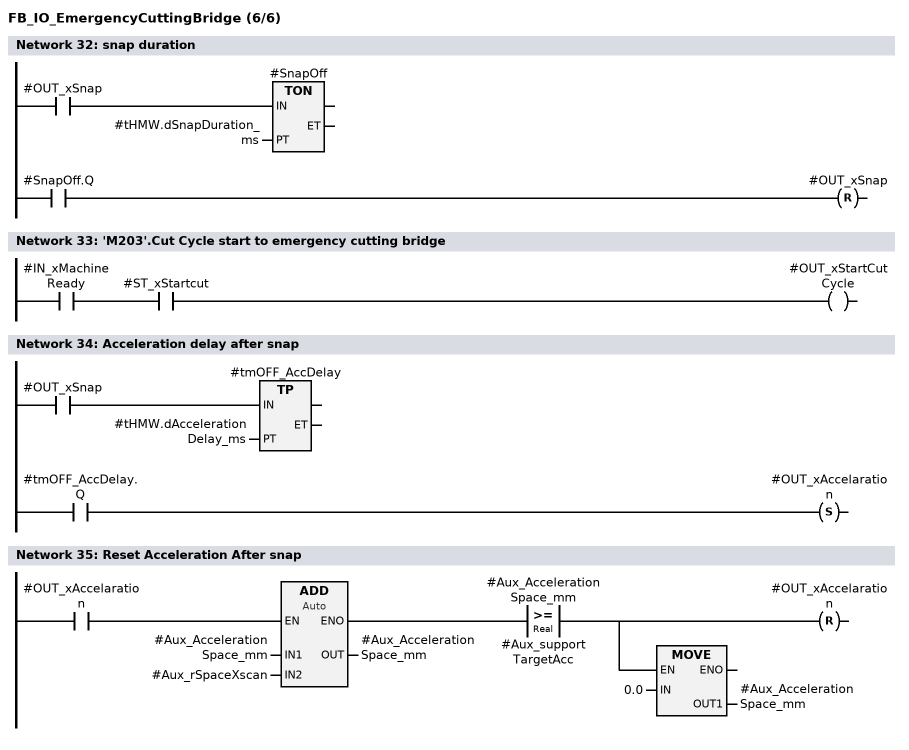
   #SnapOff(IN := #OUT_xSnap, PT := #tHMW.dSnapDuration_ms);   // TON
   IF #SnapOff.Q THEN #OUT_xSnap := FALSE; END_IF;
END_REGION

REGION Network 33: 'M203'.Cut Cycle start to emergency cutting bridge
   RUNG wire#powerrail
      Contact( #IN_xMachineReady )
      Contact( #ST_xStartcut )
      Coil( #OUT_xStartCutCycle )
   END_RUNG
   // the same network as SCL:
   #OUT_xStartCutCycle := #IN_xMachineReady AND #ST_xStartcut;
END_REGION

REGION Network 34: Acceleration delay after snap
   #tmOFF_AccDelay(IN := #OUT_xSnap, PT := #tHMW.dAccelerationDelay_ms);   // TP
   IF #tmOFF_AccDelay.Q THEN #OUT_xAccelaration := TRUE; END_IF;
END_REGION

REGION Network 35: Reset Acceleration After snap
   RUNG wire#powerrail
      Contact( #OUT_xAccelaration )
      Add(in1 := #Aux_AccelerationSpace_mm, in2 := #Aux_rSpaceXscan, out => #Aux_AccelerationSpace_mm)
      { S7_Templates := "SrcType := Real" } GE_Contact(in1 := #Aux_AccelerationSpace_mm, in2 := #Aux_supportTargetAcc)
      wire#w1
      R_Coil( #OUT_xAccelaration )
   END_RUNG
   RUNG wire#w1
      Move(in := 0.0, out1 => #Aux_AccelerationSpace_mm)
   END_RUNG
   // the same network as SCL:
   IF #OUT_xAccelaration THEN
       #Aux_AccelerationSpace_mm := #Aux_AccelerationSpace_mm + #Aux_rSpaceXscan;
   END_IF;
   #_w1 := #OUT_xAccelaration AND (#Aux_AccelerationSpace_mm >= #Aux_supportTargetAcc);
   IF #_w1 THEN
       #OUT_xAccelaration := FALSE;
       #Aux_AccelerationSpace_mm := 0.0;
   END_IF;
END_REGION
END_FUNCTION_BLOCK

// folder: 05_Reports

FUNCTION "RP_MergeToMergeMessageV2" : Void   // FC3, SCL
TITLE = RP_MergeMessage
{ S7_Optimized_Access := 'TRUE' }
AUTHOR : Cigliutt
FAMILY : RP
VERSION : 1.0
// This FC will be merge different flush buffer
   VAR_INPUT
      IN_xInit : Bool;   // Initialize the buffer container
   END_VAR
   VAR_IN_OUT
      INO_tMergeBuffer : "UDT_RP_MessageContMerge_v2";   // Merge buffer container
      INO_tMergeBuffer_1 : "UDT_RP_MessageContMerge_v2";   // Merge buffer container #1
      INO_tMergeBuffer_2 : "UDT_RP_MessageContMerge_v2";   // Merge buffer container #2
      INO_tMergeBuffer_3 : "UDT_RP_MessageContMerge_v2";   // Merge buffer container #3
      INO_tMergeBuffer_4 : "UDT_RP_MessageContMerge_v2";   // Merge buffer container #4
      INO_tMergeBuffer_5 : "UDT_RP_MessageContMerge_v2";   // Merge buffer container #5
      INO_xError : Bool;   // If =true error on flush
   END_VAR
   VAR_TEMP
      TMP_dIndex : DInt;
      TMP_dArrayNumEl : DInt;
      TMP_dtDateTime : Date_And_Time;
      TMP_dRetVal : DInt;
      TMP_dDataToCopy : DInt;
      TMP_dOldNumMex : DInt;
      TMP_dActualNumMex : DInt;
   END_VAR
BEGIN
   //Manage the initialization request. Fill to 0 the buffer and the values.
   //After that calculate the space available
   //
   #TMP_dRetVal := RD_LOC_T(#TMP_dtDateTime);

   IF #IN_xInit = true THEN

       //Initialize the values
       #INO_tMergeBuffer.dNumOfMessage := 0;
       #INO_tMergeBuffer.dMaxNumOfMessage := 0;

       //Take the number OF elements OF the array data, reset it AND set the number
       //to iDataMaxElem
       #TMP_dArrayNumEl := "GP_GetArraySize"(INO_vArray := #INO_tMergeBuffer.rgtMessages);

       #INO_tMergeBuffer.dMaxNumOfMessage := #TMP_dArrayNumEl;

       //Reset the buffer
       //

       FOR #TMP_dIndex := 0 TO #INO_tMergeBuffer.dMaxNumOfMessage - 1 DO
           #INO_tMergeBuffer.rgtMessages[#TMP_dIndex].dCodeEvent := 0;
           #INO_tMergeBuffer.rgtMessages[#TMP_dIndex].dEvent1 := 0;
           #INO_tMergeBuffer.rgtMessages[#TMP_dIndex].dEvent2 := 0;
           #INO_tMergeBuffer.rgtMessages[#TMP_dIndex].dEvent3 := 0;
           #INO_tMergeBuffer.rgtMessages[#TMP_dIndex].dEvent4 := 0;
           #INO_tMergeBuffer.rgtMessages[#TMP_dIndex].dEvent5 := 0;
           #INO_tMergeBuffer.rgtMessages[#TMP_dIndex].dEvent6 := 0;
           #INO_tMergeBuffer.rgtMessages[#TMP_dIndex].dEvent7 := 0;
           #INO_tMergeBuffer.rgtMessages[#TMP_dIndex].dEvent8 := 0;
           #INO_tMergeBuffer.rgtMessages[#TMP_dIndex].dEvent9 := 0;
           #INO_tMergeBuffer.rgtMessages[#TMP_dIndex].dEvent10 := 0;

           #INO_tMergeBuffer.rgtMessages[#TMP_dIndex].strIdent := '';
           #INO_tMergeBuffer.rgtMessages[#TMP_dIndex].dtDateTime := #TMP_dtDateTime;
       END_FOR;

       #INO_tMergeBuffer.xInitialized := true;

       RETURN;
   END_IF;

   //If we are not in initializing mode, copy the input value inside the array.
   //First of all check if the data are consistent
   //
   IF (#INO_tMergeBuffer.xInitialized = false) OR
       (#INO_tMergeBuffer_1.xInitialized = false) OR
       (#INO_tMergeBuffer_2.xInitialized = false) OR
       (#INO_tMergeBuffer_3.xInitialized = false) OR
       (#INO_tMergeBuffer_4.xInitialized = false) OR
       (#INO_tMergeBuffer_5.xInitialized = false) THEN

       #INO_xError := true;

       RETURN;
   END_IF;

   //Check if the merge buffer is free. Otherwise exit
   //
   IF (#INO_tMergeBuffer.dNumOfMessage > 0) THEN
       RETURN;
   END_IF;


   ///*********************************** FLUSH BUFFER #1

   //Check if the first flush buffer, has data inside
   IF (#INO_tMergeBuffer_1.dNumOfMessage > 0) THEN

       #TMP_dDataToCopy := #INO_tMergeBuffer_1.dNumOfMessage;

       IF (#TMP_dDataToCopy > #INO_tMergeBuffer.dMaxNumOfMessage) THEN
           #TMP_dDataToCopy := #INO_tMergeBuffer.dMaxNumOfMessage;
       END_IF;

       //Copy the data
       #TMP_dRetVal := "GP_BlockMoveStruct"(IN_iSourceIndex := 0,
                                            IN_iDestIndex := 0,
                                            IN_iCount := DINT_TO_INT(#TMP_dDataToCopy),
                                            INO_vSourceArrayStruct := #INO_tMergeBuffer_1.rgtMessages,
                                            INO_vDestArrayStruct := #INO_tMergeBuffer.rgtMessages);

       #INO_tMergeBuffer.dNumOfMessage := #TMP_dDataToCopy;

       //Check if some data is remaining. If yes, compact it on the FlushBuffer
       //
       IF (#INO_tMergeBuffer_1.dNumOfMessage - #TMP_dDataToCopy) > 0 THEN
           //Copy the data
           #TMP_dRetVal := "GP_BlockMoveStruct"(IN_iSourceIndex := DINT_TO_INT(#INO_tMergeBuffer_1.dNumOfMessage - (#INO_tMergeBuffer_1.dNumOfMessage - #TMP_dDataToCopy)),
                                                IN_iDestIndex := 0,
                                                IN_iCount := DINT_TO_INT(#INO_tMergeBuffer_1.dNumOfMessage - #TMP_dDataToCopy),
                                                INO_vSourceArrayStruct := #INO_tMergeBuffer_1.rgtMessages,
                                                INO_vDestArrayStruct := #INO_tMergeBuffer_1.rgtMessages);


       END_IF;

       #TMP_dOldNumMex := #INO_tMergeBuffer_1.dNumOfMessage;
       #TMP_dActualNumMex := #INO_tMergeBuffer_1.dNumOfMessage - #TMP_dDataToCopy;


       //Data moved, fill the remaining buffer. To increase performance, fill only the data that was used
       //
       FOR #TMP_dIndex := #TMP_dActualNumMex TO #TMP_dOldNumMex - 1 DO

           #INO_tMergeBuffer_1.rgtMessages[#TMP_dIndex].dCodeEvent := 0;
           #INO_tMergeBuffer_1.rgtMessages[#TMP_dIndex].dEvent1 := 0;
           #INO_tMergeBuffer_1.rgtMessages[#TMP_dIndex].dEvent2 := 0;
           #INO_tMergeBuffer_1.rgtMessages[#TMP_dIndex].dEvent3 := 0;
           #INO_tMergeBuffer_1.rgtMessages[#TMP_dIndex].dEvent4 := 0;
           #INO_tMergeBuffer_1.rgtMessages[#TMP_dIndex].dEvent5 := 0;
           #INO_tMergeBuffer_1.rgtMessages[#TMP_dIndex].dEvent6 := 0;
           #INO_tMergeBuffer_1.rgtMessages[#TMP_dIndex].dEvent7 := 0;
           #INO_tMergeBuffer_1.rgtMessages[#TMP_dIndex].dEvent8 := 0;
           #INO_tMergeBuffer_1.rgtMessages[#TMP_dIndex].dEvent9 := 0;
           #INO_tMergeBuffer_1.rgtMessages[#TMP_dIndex].dEvent10 := 0;

           #INO_tMergeBuffer_1.rgtMessages[#TMP_dIndex].strIdent := '';
           #INO_tMergeBuffer_1.rgtMessages[#TMP_dIndex].dtDateTime := #TMP_dtDateTime;
       END_FOR;

       #INO_tMergeBuffer_1.dNumOfMessage := #TMP_dActualNumMex;

   END_IF;


   ///*********************************** FLUSH BUFFER #2

   //Check if the first flush buffer, has data inside
   IF (#INO_tMergeBuffer_2.dNumOfMessage > 0) AND (#INO_tMergeBuffer.dNumOfMessage < #INO_tMergeBuffer.dMaxNumOfMessage) THEN

       #TMP_dDataToCopy := #INO_tMergeBuffer_2.dNumOfMessage;

       IF (#TMP_dDataToCopy + #INO_tMergeBuffer.dNumOfMessage > #INO_tMergeBuffer.dMaxNumOfMessage) THEN
           #TMP_dDataToCopy := #INO_tMergeBuffer.dMaxNumOfMessage - #INO_tMergeBuffer.dNumOfMessage;
       END_IF;

       //Copy the data
       #TMP_dRetVal := "GP_BlockMoveStruct"(IN_iSourceIndex := 0,
                                            IN_iDestIndex := DINT_TO_INT(#INO_tMergeBuffer.dNumOfMessage),
                                            IN_iCount := DINT_TO_INT(#TMP_dDataToCopy),
                                            INO_vSourceArrayStruct := #INO_tMergeBuffer_2.rgtMessages,
                                            INO_vDestArrayStruct := #INO_tMergeBuffer.rgtMessages);

       #INO_tMergeBuffer.dNumOfMessage := #INO_tMergeBuffer.dNumOfMessage + #TMP_dDataToCopy;

       //Check if some data is remaining. If yes, compact it on the FlushBuffer
       //
       IF (#INO_tMergeBuffer_2.dNumOfMessage - #TMP_dDataToCopy) > 0 THEN
           //Copy the data
           #TMP_dRetVal := "GP_BlockMoveStruct"(IN_iSourceIndex := DINT_TO_INT(#INO_tMergeBuffer_2.dNumOfMessage - (#INO_tMergeBuffer_2.dNumOfMessage - #TMP_dDataToCopy)),
                                                IN_iDestIndex := 0,
                                                IN_iCount := DINT_TO_INT(#INO_tMergeBuffer_2.dNumOfMessage - #TMP_dDataToCopy),
                                                INO_vSourceArrayStruct := #INO_tMergeBuffer_2.rgtMessages,
                                                INO_vDestArrayStruct := #INO_tMergeBuffer_2.rgtMessages);


       END_IF;

       #TMP_dOldNumMex := #INO_tMergeBuffer_2.dNumOfMessage;
       #TMP_dActualNumMex := #INO_tMergeBuffer_2.dNumOfMessage - #TMP_dDataToCopy;



       //Data moved, fill the remaining buffer. To increase performance, fill only the data that was used
       //
       FOR #TMP_dIndex := #TMP_dActualNumMex TO #TMP_dOldNumMex - 1 DO

           #INO_tMergeBuffer_2.rgtMessages[#TMP_dIndex].dCodeEvent := 0;
           #INO_tMergeBuffer_2.rgtMessages[#TMP_dIndex].dEvent1 := 0;
           #INO_tMergeBuffer_2.rgtMessages[#TMP_dIndex].dEvent2 := 0;
           #INO_tMergeBuffer_2.rgtMessages[#TMP_dIndex].dEvent3 := 0;
           #INO_tMergeBuffer_2.rgtMessages[#TMP_dIndex].dEvent4 := 0;
           #INO_tMergeBuffer_2.rgtMessages[#TMP_dIndex].dEvent5 := 0;
           #INO_tMergeBuffer_2.rgtMessages[#TMP_dIndex].dEvent6 := 0;
           #INO_tMergeBuffer_2.rgtMessages[#TMP_dIndex].dEvent7 := 0;
           #INO_tMergeBuffer_2.rgtMessages[#TMP_dIndex].dEvent8 := 0;
           #INO_tMergeBuffer_2.rgtMessages[#TMP_dIndex].dEvent9 := 0;
           #INO_tMergeBuffer_2.rgtMessages[#TMP_dIndex].dEvent10 := 0;
           #INO_tMergeBuffer_2.rgtMessages[#TMP_dIndex].strIdent := '';

           #INO_tMergeBuffer_2.rgtMessages[#TMP_dIndex].dtDateTime := #TMP_dtDateTime;
       END_FOR;

       #INO_tMergeBuffer_2.dNumOfMessage := #TMP_dActualNumMex;
   END_IF;


   ///*********************************** FLUSH BUFFER #3


   //Check if the first flush buffer, has data inside
   IF (#INO_tMergeBuffer_3.dNumOfMessage > 0) AND (#INO_tMergeBuffer.dNumOfMessage < #INO_tMergeBuffer.dMaxNumOfMessage) THEN

       #TMP_dDataToCopy := #INO_tMergeBuffer_3.dNumOfMessage;

       IF (#TMP_dDataToCopy + #INO_tMergeBuffer.dNumOfMessage > #INO_tMergeBuffer.dMaxNumOfMessage) THEN
           #TMP_dDataToCopy := #INO_tMergeBuffer.dMaxNumOfMessage - #INO_tMergeBuffer.dNumOfMessage;
       END_IF;

       //Copy the data
       #TMP_dRetVal := "GP_BlockMoveStruct"(IN_iSourceIndex := 0,
                                            IN_iDestIndex := DINT_TO_INT(#INO_tMergeBuffer.dNumOfMessage),
                                            IN_iCount := DINT_TO_INT(#TMP_dDataToCopy),
                                            INO_vSourceArrayStruct := #INO_tMergeBuffer_3.rgtMessages,
                                            INO_vDestArrayStruct := #INO_tMergeBuffer.rgtMessages);

       #INO_tMergeBuffer.dNumOfMessage := #INO_tMergeBuffer.dNumOfMessage + #TMP_dDataToCopy;

       //Check if some data is remaining. If yes, compact it on the FlushBuffer
       //
       IF (#INO_tMergeBuffer_3.dNumOfMessage - #TMP_dDataToCopy) > 0 THEN
           //Copy the data
           #TMP_dRetVal := "GP_BlockMoveStruct"(IN_iSourceIndex := DINT_TO_INT(#INO_tMergeBuffer_3.dNumOfMessage - (#INO_tMergeBuffer_3.dNumOfMessage - #TMP_dDataToCopy)),
                                                IN_iDestIndex := 0,
                                                IN_iCount := DINT_TO_INT(#INO_tMergeBuffer_3.dNumOfMessage - #TMP_dDataToCopy),
                                                INO_vSourceArrayStruct := #INO_tMergeBuffer_3.rgtMessages,
                                                INO_vDestArrayStruct := #INO_tMergeBuffer_3.rgtMessages);


       END_IF;

       #TMP_dOldNumMex := #INO_tMergeBuffer_3.dNumOfMessage;
       #TMP_dActualNumMex := #INO_tMergeBuffer_3.dNumOfMessage - #TMP_dDataToCopy;


       //Data moved, fill the remaining buffer. To increase performance, fill only the data that was used
       //
       FOR #TMP_dIndex := #TMP_dActualNumMex TO #TMP_dOldNumMex - 1 DO

           #INO_tMergeBuffer_3.rgtMessages[#TMP_dIndex].dCodeEvent := 0;
           #INO_tMergeBuffer_3.rgtMessages[#TMP_dIndex].dEvent1 := 0;
           #INO_tMergeBuffer_3.rgtMessages[#TMP_dIndex].dEvent2 := 0;
           #INO_tMergeBuffer_3.rgtMessages[#TMP_dIndex].dEvent3 := 0;
           #INO_tMergeBuffer_3.rgtMessages[#TMP_dIndex].dEvent4 := 0;
           #INO_tMergeBuffer_3.rgtMessages[#TMP_dIndex].dEvent5 := 0;
           #INO_tMergeBuffer_3.rgtMessages[#TMP_dIndex].dEvent6 := 0;
           #INO_tMergeBuffer_3.rgtMessages[#TMP_dIndex].dEvent7 := 0;
           #INO_tMergeBuffer_3.rgtMessages[#TMP_dIndex].dEvent8 := 0;
           #INO_tMergeBuffer_3.rgtMessages[#TMP_dIndex].dEvent9 := 0;
           #INO_tMergeBuffer_3.rgtMessages[#TMP_dIndex].dEvent10 := 0;
           #INO_tMergeBuffer_3.rgtMessages[#TMP_dIndex].strIdent := '';

           #INO_tMergeBuffer_3.rgtMessages[#TMP_dIndex].dtDateTime := #TMP_dtDateTime;
       END_FOR;

       #INO_tMergeBuffer_3.dNumOfMessage := #TMP_dActualNumMex;


   END_IF;


   ///*********************************** FLUSH BUFFER #4


   //Check if the first flush buffer, has data inside
   IF (#INO_tMergeBuffer_4.dNumOfMessage > 0) AND (#INO_tMergeBuffer.dNumOfMessage < #INO_tMergeBuffer.dMaxNumOfMessage) THEN

       #TMP_dDataToCopy := #INO_tMergeBuffer_4.dNumOfMessage;

       IF (#TMP_dDataToCopy + #INO_tMergeBuffer.dNumOfMessage > #INO_tMergeBuffer.dMaxNumOfMessage) THEN
           #TMP_dDataToCopy := #INO_tMergeBuffer.dMaxNumOfMessage - #INO_tMergeBuffer.dNumOfMessage;
       END_IF;

       //Copy the data
       #TMP_dRetVal := "GP_BlockMoveStruct"(IN_iSourceIndex := 0,
                                            IN_iDestIndex := DINT_TO_INT(#INO_tMergeBuffer.dNumOfMessage),
                                            IN_iCount := DINT_TO_INT(#TMP_dDataToCopy),
                                            INO_vSourceArrayStruct := #INO_tMergeBuffer_4.rgtMessages,
                                            INO_vDestArrayStruct := #INO_tMergeBuffer.rgtMessages);

       #INO_tMergeBuffer.dNumOfMessage := #INO_tMergeBuffer.dNumOfMessage + #TMP_dDataToCopy;

       //Check if some data is remaining. If yes, compact it on the FlushBuffer
       //
       IF (#INO_tMergeBuffer_4.dNumOfMessage - #TMP_dDataToCopy) > 0 THEN
           //Copy the data
           #TMP_dRetVal := "GP_BlockMoveStruct"(IN_iSourceIndex := DINT_TO_INT(#INO_tMergeBuffer_4.dNumOfMessage - (#INO_tMergeBuffer_4.dNumOfMessage - #TMP_dDataToCopy)),
                                                IN_iDestIndex := 0,
                                                IN_iCount := DINT_TO_INT(#INO_tMergeBuffer_4.dNumOfMessage - #TMP_dDataToCopy),
                                                INO_vSourceArrayStruct := #INO_tMergeBuffer_4.rgtMessages,
                                                INO_vDestArrayStruct := #INO_tMergeBuffer_4.rgtMessages);


       END_IF;

       #TMP_dOldNumMex := #INO_tMergeBuffer_4.dNumOfMessage;
       #TMP_dActualNumMex := #INO_tMergeBuffer_4.dNumOfMessage - #TMP_dDataToCopy;


       //Data moved, fill the remaining buffer. To increase performance, fill only the data that was used
       //
       FOR #TMP_dIndex := #TMP_dActualNumMex TO #TMP_dOldNumMex - 1 DO

           #INO_tMergeBuffer_4.rgtMessages[#TMP_dIndex].dCodeEvent := 0;
           #INO_tMergeBuffer_4.rgtMessages[#TMP_dIndex].dEvent1 := 0;
           #INO_tMergeBuffer_4.rgtMessages[#TMP_dIndex].dEvent2 := 0;
           #INO_tMergeBuffer_4.rgtMessages[#TMP_dIndex].dEvent3 := 0;
           #INO_tMergeBuffer_4.rgtMessages[#TMP_dIndex].dEvent4 := 0;
           #INO_tMergeBuffer_4.rgtMessages[#TMP_dIndex].dEvent5 := 0;
           #INO_tMergeBuffer_4.rgtMessages[#TMP_dIndex].dEvent6 := 0;
           #INO_tMergeBuffer_4.rgtMessages[#TMP_dIndex].dEvent7 := 0;
           #INO_tMergeBuffer_4.rgtMessages[#TMP_dIndex].dEvent8 := 0;
           #INO_tMergeBuffer_4.rgtMessages[#TMP_dIndex].dEvent9 := 0;
           #INO_tMergeBuffer_4.rgtMessages[#TMP_dIndex].dEvent10 := 0;
           #INO_tMergeBuffer_4.rgtMessages[#TMP_dIndex].strIdent := '';

           #INO_tMergeBuffer_4.rgtMessages[#TMP_dIndex].dtDateTime := #TMP_dtDateTime;
       END_FOR;

       #INO_tMergeBuffer_4.dNumOfMessage := #TMP_dActualNumMex;


   END_IF;


   ///*********************************** FLUSH BUFFER #5


   //Check if the first flush buffer, has data inside
   IF (#INO_tMergeBuffer_5.dNumOfMessage > 0) AND (#INO_tMergeBuffer.dNumOfMessage < #INO_tMergeBuffer.dMaxNumOfMessage) THEN

       #TMP_dDataToCopy := #INO_tMergeBuffer_5.dNumOfMessage;

       IF (#TMP_dDataToCopy + #INO_tMergeBuffer.dNumOfMessage > #INO_tMergeBuffer.dMaxNumOfMessage) THEN
           #TMP_dDataToCopy := #INO_tMergeBuffer.dMaxNumOfMessage - #INO_tMergeBuffer.dNumOfMessage;
       END_IF;

       //Copy the data
       #TMP_dRetVal := "GP_BlockMoveStruct"(IN_iSourceIndex := 0,
                                            IN_iDestIndex := DINT_TO_INT(#INO_tMergeBuffer.dNumOfMessage),
                                            IN_iCount := DINT_TO_INT(#TMP_dDataToCopy),
                                            INO_vSourceArrayStruct := #INO_tMergeBuffer_5.rgtMessages,
                                            INO_vDestArrayStruct := #INO_tMergeBuffer.rgtMessages);

       #INO_tMergeBuffer.dNumOfMessage := #INO_tMergeBuffer.dNumOfMessage + #TMP_dDataToCopy;

       //Check if some data is remaining. If yes, compact it on the FlushBuffer
       //
       IF (#INO_tMergeBuffer_5.dNumOfMessage - #TMP_dDataToCopy) > 0 THEN
           //Copy the data
           #TMP_dRetVal := "GP_BlockMoveStruct"(IN_iSourceIndex := DINT_TO_INT(#INO_tMergeBuffer_5.dNumOfMessage - (#INO_tMergeBuffer_5.dNumOfMessage - #TMP_dDataToCopy)),
                                                IN_iDestIndex := 0,
                                                IN_iCount := DINT_TO_INT(#INO_tMergeBuffer_5.dNumOfMessage - #TMP_dDataToCopy),
                                                INO_vSourceArrayStruct := #INO_tMergeBuffer_5.rgtMessages,
                                                INO_vDestArrayStruct := #INO_tMergeBuffer_5.rgtMessages);


       END_IF;

       #TMP_dOldNumMex := #INO_tMergeBuffer_5.dNumOfMessage;
       #TMP_dActualNumMex := #INO_tMergeBuffer_5.dNumOfMessage - #TMP_dDataToCopy;

       //Data moved, fill the remaining buffer. To increase performance, fill only the data that was used
       //
       FOR #TMP_dIndex := #TMP_dActualNumMex TO #TMP_dOldNumMex - 1 DO

           #INO_tMergeBuffer_5.rgtMessages[#TMP_dIndex].dCodeEvent := 0;
           #INO_tMergeBuffer_5.rgtMessages[#TMP_dIndex].dEvent1 := 0;
           #INO_tMergeBuffer_5.rgtMessages[#TMP_dIndex].dEvent2 := 0;
           #INO_tMergeBuffer_5.rgtMessages[#TMP_dIndex].dEvent3 := 0;
           #INO_tMergeBuffer_5.rgtMessages[#TMP_dIndex].dEvent4 := 0;
           #INO_tMergeBuffer_5.rgtMessages[#TMP_dIndex].dEvent5 := 0;
           #INO_tMergeBuffer_5.rgtMessages[#TMP_dIndex].dEvent6 := 0;
           #INO_tMergeBuffer_5.rgtMessages[#TMP_dIndex].dEvent7 := 0;
           #INO_tMergeBuffer_5.rgtMessages[#TMP_dIndex].dEvent8 := 0;
           #INO_tMergeBuffer_5.rgtMessages[#TMP_dIndex].dEvent9 := 0;
           #INO_tMergeBuffer_5.rgtMessages[#TMP_dIndex].dEvent10 := 0;
           #INO_tMergeBuffer_5.rgtMessages[#TMP_dIndex].strIdent := '';

           #INO_tMergeBuffer_5.rgtMessages[#TMP_dIndex].dtDateTime := #TMP_dtDateTime;
       END_FOR;

       #INO_tMergeBuffer_5.dNumOfMessage := #TMP_dActualNumMex;


   END_IF;
END_FUNCTION

FUNCTION "RP_OB_TaskSlowToOpt" : Void   // FC4, LAD
{ S7_Optimized_Access := 'TRUE' }
VERSION : 0.1
   VAR_INPUT
      IN_xFirstScan : Bool;
   END_VAR
   VAR_TEMP
      TMP_xError : Bool;
   END_VAR
BEGIN

REGION Network 1
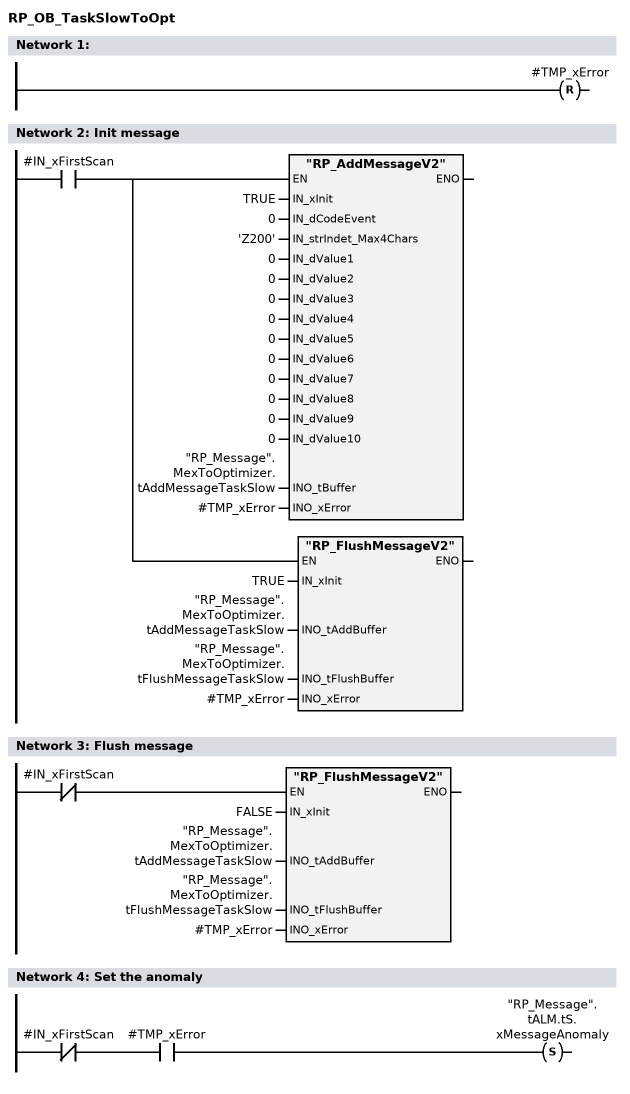
   RUNG wire#powerrail
      R_Coil( #TMP_xError )
   END_RUNG
   // the same network as SCL:
   #TMP_xError := FALSE;
END_REGION

REGION Network 2: Init message
   RUNG wire#powerrail
      Contact( #IN_xFirstScan )
      wire#w1
      "RP_AddMessageV2"(IN_xInit := TRUE, IN_dCodeEvent := 0, IN_strIndet_Max4Chars := 'Z200', IN_dValue1 := 0, IN_dValue2 := 0, IN_dValue3 := 0, IN_dValue4 := 0, IN_dValue5 := 0, IN_dValue6 := 0, IN_dValue7 := 0, IN_dValue8 := 0, IN_dValue9 := 0, IN_dValue10 := 0, INO_tBuffer := "RP_Message".MexToOptimizer.tAddMessageTaskSlow, INO_xError := #TMP_xError)
   END_RUNG
   RUNG wire#w1
      "RP_FlushMessageV2"(IN_xInit := TRUE, INO_tAddBuffer := "RP_Message".MexToOptimizer.tAddMessageTaskSlow, INO_tFlushBuffer := "RP_Message".MexToOptimizer.tFlushMessageTaskSlow, INO_xError := #TMP_xError)
   END_RUNG
   // the same network as SCL:
   IF #IN_xFirstScan THEN
       "RP_AddMessageV2"(IN_xInit := TRUE,
                         IN_dCodeEvent := 0,
                         IN_strIndet_Max4Chars := 'Z200',
                         IN_dValue1 := 0,
                         IN_dValue2 := 0,
                         IN_dValue3 := 0,
                         IN_dValue4 := 0,
                         IN_dValue5 := 0,
                         IN_dValue6 := 0,
                         IN_dValue7 := 0,
                         IN_dValue8 := 0,
                         IN_dValue9 := 0,
                         IN_dValue10 := 0,
                         INO_tBuffer := "RP_Message".MexToOptimizer.tAddMessageTaskSlow,
                         INO_xError := #TMP_xError);
       "RP_FlushMessageV2"(IN_xInit := TRUE,
                           INO_tAddBuffer := "RP_Message".MexToOptimizer.tAddMessageTaskSlow,
                           INO_tFlushBuffer := "RP_Message".MexToOptimizer.tFlushMessageTaskSlow,
                           INO_xError := #TMP_xError);
   END_IF;
END_REGION

REGION Network 3: Flush message
   RUNG wire#powerrail
      I_Contact( #IN_xFirstScan )
      "RP_FlushMessageV2"(IN_xInit := FALSE, INO_tAddBuffer := "RP_Message".MexToOptimizer.tAddMessageTaskSlow, INO_tFlushBuffer := "RP_Message".MexToOptimizer.tFlushMessageTaskSlow, INO_xError := #TMP_xError)
   END_RUNG
   // the same network as SCL:
   IF NOT #IN_xFirstScan THEN
       "RP_FlushMessageV2"(IN_xInit := FALSE,
                           INO_tAddBuffer := "RP_Message".MexToOptimizer.tAddMessageTaskSlow,
                           INO_tFlushBuffer := "RP_Message".MexToOptimizer.tFlushMessageTaskSlow,
                           INO_xError := #TMP_xError);
   END_IF;
END_REGION

REGION Network 4: Set the anomaly
   RUNG wire#powerrail
      I_Contact( #IN_xFirstScan )
      Contact( #TMP_xError )
      S_Coil( "RP_Message".tALM.tS.xMessageAnomaly )
   END_RUNG
   // the same network as SCL:
   IF NOT #IN_xFirstScan AND #TMP_xError THEN "RP_Message".tALM.tS.xMessageAnomaly := TRUE; END_IF;
END_REGION
END_FUNCTION

FUNCTION "RP_OB_TaskMediumFromOpt" : Void   // FC5, LAD
{ S7_Optimized_Access := 'TRUE' }
VERSION : 0.1
   VAR_INPUT
      IN_xFirstScan : Bool;
   END_VAR
   VAR_TEMP
      TMP_xError : Bool;
   END_VAR
BEGIN

REGION Network 1
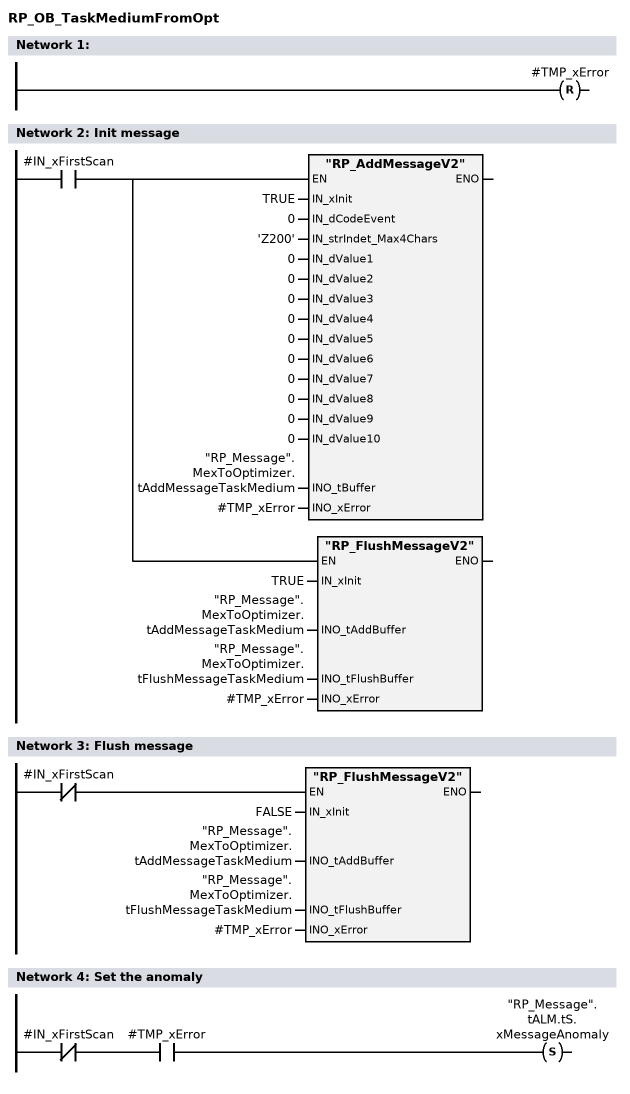
   RUNG wire#powerrail
      R_Coil( #TMP_xError )
   END_RUNG
   // the same network as SCL:
   #TMP_xError := FALSE;
END_REGION

REGION Network 2: Init message
   RUNG wire#powerrail
      Contact( #IN_xFirstScan )
      wire#w1
      "RP_AddMessageV2"(IN_xInit := TRUE, IN_dCodeEvent := 0, IN_strIndet_Max4Chars := 'Z200', IN_dValue1 := 0, IN_dValue2 := 0, IN_dValue3 := 0, IN_dValue4 := 0, IN_dValue5 := 0, IN_dValue6 := 0, IN_dValue7 := 0, IN_dValue8 := 0, IN_dValue9 := 0, IN_dValue10 := 0, INO_tBuffer := "RP_Message".MexToOptimizer.tAddMessageTaskMedium, INO_xError := #TMP_xError)
   END_RUNG
   RUNG wire#w1
      "RP_FlushMessageV2"(IN_xInit := TRUE, INO_tAddBuffer := "RP_Message".MexToOptimizer.tAddMessageTaskMedium, INO_tFlushBuffer := "RP_Message".MexToOptimizer.tFlushMessageTaskMedium, INO_xError := #TMP_xError)
   END_RUNG
   // the same network as SCL:
   IF #IN_xFirstScan THEN
       "RP_AddMessageV2"(IN_xInit := TRUE,
                         IN_dCodeEvent := 0,
                         IN_strIndet_Max4Chars := 'Z200',
                         IN_dValue1 := 0,
                         IN_dValue2 := 0,
                         IN_dValue3 := 0,
                         IN_dValue4 := 0,
                         IN_dValue5 := 0,
                         IN_dValue6 := 0,
                         IN_dValue7 := 0,
                         IN_dValue8 := 0,
                         IN_dValue9 := 0,
                         IN_dValue10 := 0,
                         INO_tBuffer := "RP_Message".MexToOptimizer.tAddMessageTaskMedium,
                         INO_xError := #TMP_xError);
       "RP_FlushMessageV2"(IN_xInit := TRUE,
                           INO_tAddBuffer := "RP_Message".MexToOptimizer.tAddMessageTaskMedium,
                           INO_tFlushBuffer := "RP_Message".MexToOptimizer.tFlushMessageTaskMedium,
                           INO_xError := #TMP_xError);
   END_IF;
END_REGION

REGION Network 3: Flush message
   RUNG wire#powerrail
      I_Contact( #IN_xFirstScan )
      "RP_FlushMessageV2"(IN_xInit := FALSE, INO_tAddBuffer := "RP_Message".MexToOptimizer.tAddMessageTaskMedium, INO_tFlushBuffer := "RP_Message".MexToOptimizer.tFlushMessageTaskMedium, INO_xError := #TMP_xError)
   END_RUNG
   // the same network as SCL:
   IF NOT #IN_xFirstScan THEN
       "RP_FlushMessageV2"(IN_xInit := FALSE,
                           INO_tAddBuffer := "RP_Message".MexToOptimizer.tAddMessageTaskMedium,
                           INO_tFlushBuffer := "RP_Message".MexToOptimizer.tFlushMessageTaskMedium,
                           INO_xError := #TMP_xError);
   END_IF;
END_REGION

REGION Network 4: Set the anomaly
   RUNG wire#powerrail
      I_Contact( #IN_xFirstScan )
      Contact( #TMP_xError )
      S_Coil( "RP_Message".tALM.tS.xMessageAnomaly )
   END_RUNG
   // the same network as SCL:
   IF NOT #IN_xFirstScan AND #TMP_xError THEN "RP_Message".tALM.tS.xMessageAnomaly := TRUE; END_IF;
END_REGION
END_FUNCTION

FUNCTION "RP_OB_TaskMediumToOpt" : Void   // FC6, LAD
{ S7_Optimized_Access := 'TRUE' }
VERSION : 0.1
   VAR_INPUT
      IN_xFirstScan : Bool;
   END_VAR
   VAR_TEMP
      TMP_xError : Bool;
   END_VAR
BEGIN

REGION Network 1
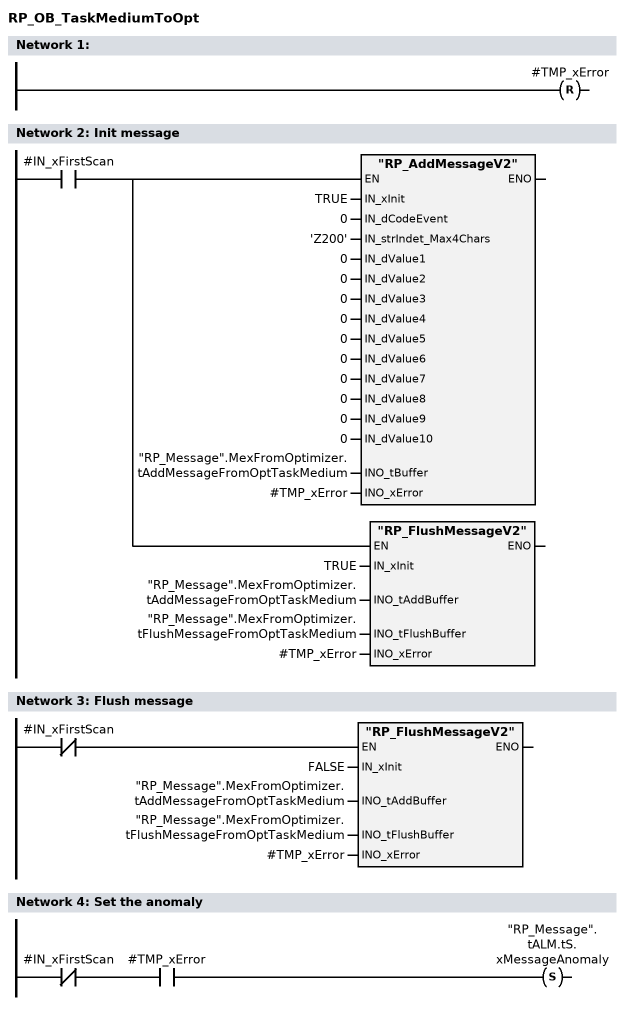
   RUNG wire#powerrail
      R_Coil( #TMP_xError )
   END_RUNG
   // the same network as SCL:
   #TMP_xError := FALSE;
END_REGION

REGION Network 2: Init message
   RUNG wire#powerrail
      Contact( #IN_xFirstScan )
      wire#w1
      "RP_AddMessageV2"(IN_xInit := TRUE, IN_dCodeEvent := 0, IN_strIndet_Max4Chars := 'Z200', IN_dValue1 := 0, IN_dValue2 := 0, IN_dValue3 := 0, IN_dValue4 := 0, IN_dValue5 := 0, IN_dValue6 := 0, IN_dValue7 := 0, IN_dValue8 := 0, IN_dValue9 := 0, IN_dValue10 := 0, INO_tBuffer := "RP_Message".MexFromOptimizer.tAddMessageFromOptTaskMedium, INO_xError := #TMP_xError)
   END_RUNG
   RUNG wire#w1
      "RP_FlushMessageV2"(IN_xInit := TRUE, INO_tAddBuffer := "RP_Message".MexFromOptimizer.tAddMessageFromOptTaskMedium, INO_tFlushBuffer := "RP_Message".MexFromOptimizer.tFlushMessageFromOptTaskMedium, INO_xError := #TMP_xError)
   END_RUNG
   // the same network as SCL:
   IF #IN_xFirstScan THEN
       "RP_AddMessageV2"(IN_xInit := TRUE,
                         IN_dCodeEvent := 0,
                         IN_strIndet_Max4Chars := 'Z200',
                         IN_dValue1 := 0,
                         IN_dValue2 := 0,
                         IN_dValue3 := 0,
                         IN_dValue4 := 0,
                         IN_dValue5 := 0,
                         IN_dValue6 := 0,
                         IN_dValue7 := 0,
                         IN_dValue8 := 0,
                         IN_dValue9 := 0,
                         IN_dValue10 := 0,
                         INO_tBuffer := "RP_Message".MexFromOptimizer.tAddMessageFromOptTaskMedium,
                         INO_xError := #TMP_xError);
       "RP_FlushMessageV2"(IN_xInit := TRUE,
                           INO_tAddBuffer := "RP_Message".MexFromOptimizer.tAddMessageFromOptTaskMedium,
                           INO_tFlushBuffer := "RP_Message".MexFromOptimizer.tFlushMessageFromOptTaskMedium,
                           INO_xError := #TMP_xError);
   END_IF;
END_REGION

REGION Network 3: Flush message
   RUNG wire#powerrail
      I_Contact( #IN_xFirstScan )
      "RP_FlushMessageV2"(IN_xInit := FALSE, INO_tAddBuffer := "RP_Message".MexFromOptimizer.tAddMessageFromOptTaskMedium, INO_tFlushBuffer := "RP_Message".MexFromOptimizer.tFlushMessageFromOptTaskMedium, INO_xError := #TMP_xError)
   END_RUNG
   // the same network as SCL:
   IF NOT #IN_xFirstScan THEN
       "RP_FlushMessageV2"(IN_xInit := FALSE,
                           INO_tAddBuffer := "RP_Message".MexFromOptimizer.tAddMessageFromOptTaskMedium,
                           INO_tFlushBuffer := "RP_Message".MexFromOptimizer.tFlushMessageFromOptTaskMedium,
                           INO_xError := #TMP_xError);
   END_IF;
END_REGION

REGION Network 4: Set the anomaly
   RUNG wire#powerrail
      I_Contact( #IN_xFirstScan )
      Contact( #TMP_xError )
      S_Coil( "RP_Message".tALM.tS.xMessageAnomaly )
   END_RUNG
   // the same network as SCL:
   IF NOT #IN_xFirstScan AND #TMP_xError THEN "RP_Message".tALM.tS.xMessageAnomaly := TRUE; END_IF;
END_REGION
END_FUNCTION

FUNCTION "RP_OB_TaskFastToOpt" : Void   // FC18, LAD
{ S7_Optimized_Access := 'TRUE' }
VERSION : 0.1
   VAR_INPUT
      IN_xFirstScan : Bool;
   END_VAR
   VAR_TEMP
      TMP_xError : Bool;
   END_VAR
BEGIN

REGION Network 1
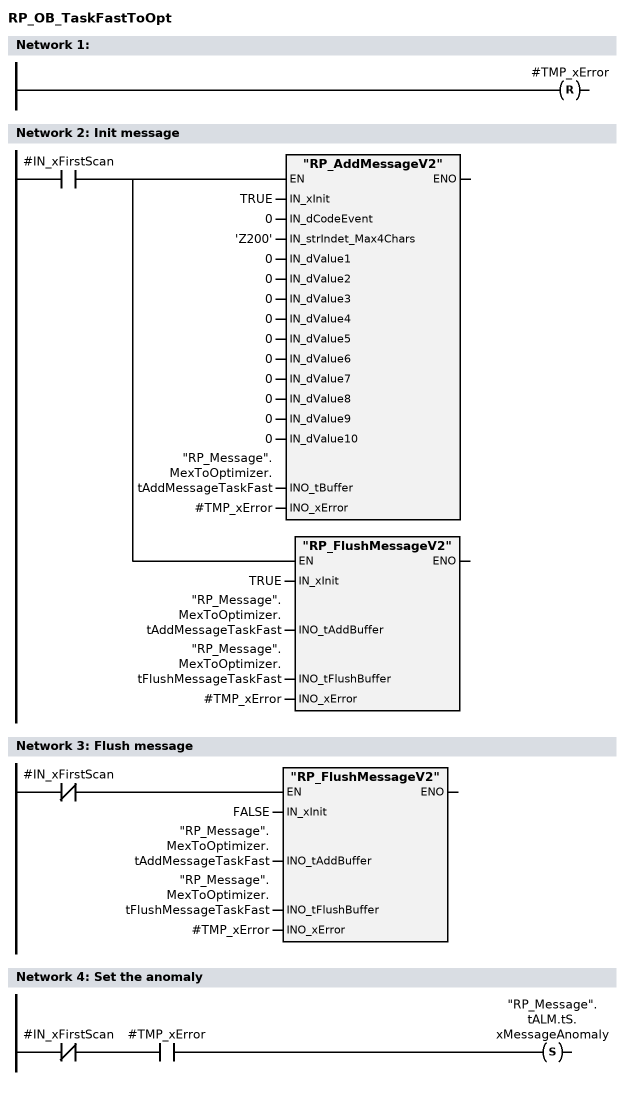
   RUNG wire#powerrail
      R_Coil( #TMP_xError )
   END_RUNG
   // the same network as SCL:
   #TMP_xError := FALSE;
END_REGION

REGION Network 2: Init message
   RUNG wire#powerrail
      Contact( #IN_xFirstScan )
      wire#w1
      "RP_AddMessageV2"(IN_xInit := TRUE, IN_dCodeEvent := 0, IN_strIndet_Max4Chars := 'Z200', IN_dValue1 := 0, IN_dValue2 := 0, IN_dValue3 := 0, IN_dValue4 := 0, IN_dValue5 := 0, IN_dValue6 := 0, IN_dValue7 := 0, IN_dValue8 := 0, IN_dValue9 := 0, IN_dValue10 := 0, INO_tBuffer := "RP_Message".MexToOptimizer.tAddMessageTaskFast, INO_xError := #TMP_xError)
   END_RUNG
   RUNG wire#w1
      "RP_FlushMessageV2"(IN_xInit := TRUE, INO_tAddBuffer := "RP_Message".MexToOptimizer.tAddMessageTaskFast, INO_tFlushBuffer := "RP_Message".MexToOptimizer.tFlushMessageTaskFast, INO_xError := #TMP_xError)
   END_RUNG
   // the same network as SCL:
   IF #IN_xFirstScan THEN
       "RP_AddMessageV2"(IN_xInit := TRUE,
                         IN_dCodeEvent := 0,
                         IN_strIndet_Max4Chars := 'Z200',
                         IN_dValue1 := 0,
                         IN_dValue2 := 0,
                         IN_dValue3 := 0,
                         IN_dValue4 := 0,
                         IN_dValue5 := 0,
                         IN_dValue6 := 0,
                         IN_dValue7 := 0,
                         IN_dValue8 := 0,
                         IN_dValue9 := 0,
                         IN_dValue10 := 0,
                         INO_tBuffer := "RP_Message".MexToOptimizer.tAddMessageTaskFast,
                         INO_xError := #TMP_xError);
       "RP_FlushMessageV2"(IN_xInit := TRUE,
                           INO_tAddBuffer := "RP_Message".MexToOptimizer.tAddMessageTaskFast,
                           INO_tFlushBuffer := "RP_Message".MexToOptimizer.tFlushMessageTaskFast,
                           INO_xError := #TMP_xError);
   END_IF;
END_REGION

REGION Network 3: Flush message
   RUNG wire#powerrail
      I_Contact( #IN_xFirstScan )
      "RP_FlushMessageV2"(IN_xInit := FALSE, INO_tAddBuffer := "RP_Message".MexToOptimizer.tAddMessageTaskFast, INO_tFlushBuffer := "RP_Message".MexToOptimizer.tFlushMessageTaskFast, INO_xError := #TMP_xError)
   END_RUNG
   // the same network as SCL:
   IF NOT #IN_xFirstScan THEN
       "RP_FlushMessageV2"(IN_xInit := FALSE,
                           INO_tAddBuffer := "RP_Message".MexToOptimizer.tAddMessageTaskFast,
                           INO_tFlushBuffer := "RP_Message".MexToOptimizer.tFlushMessageTaskFast,
                           INO_xError := #TMP_xError);
   END_IF;
END_REGION

REGION Network 4: Set the anomaly
   RUNG wire#powerrail
      I_Contact( #IN_xFirstScan )
      Contact( #TMP_xError )
      S_Coil( "RP_Message".tALM.tS.xMessageAnomaly )
   END_RUNG
   // the same network as SCL:
   IF NOT #IN_xFirstScan AND #TMP_xError THEN "RP_Message".tALM.tS.xMessageAnomaly := TRUE; END_IF;
END_REGION
END_FUNCTION

FUNCTION "RP_OB_TaskMainToOpt" : Void   // FC19, LAD
{ S7_Optimized_Access := 'TRUE' }
VERSION : 0.1
   VAR_INPUT
      IN_xFirstScan : Bool;
   END_VAR
   VAR_TEMP
      TMP_xError : Bool;
      TMP_iRet : Int;
      TMP_dwValue : DWord;
   END_VAR
BEGIN

REGION Network 1: Reset temporary
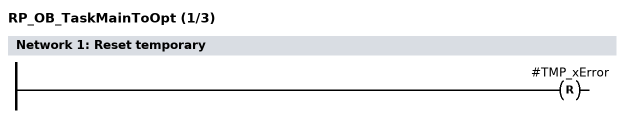
   RUNG wire#powerrail
      R_Coil( #TMP_xError )
   END_RUNG
   // the same network as SCL:
   #TMP_xError := FALSE;
END_REGION

REGION Network 2 (SCL): Reset alarms
   IF "Z201".tmOFF_ResetAlarm.OUT_xDone THEN

       #TMP_dwValue := 0;

       SCATTER(IN:=#TMP_dwValue,
               OUT=>"RP_Message".tALM.tS);

       SCATTER(IN:=#TMP_dwValue,
               OUT=>"RP_Message".tALM.tF);

       SCATTER(IN:=#TMP_dwValue,
               OUT=>"RP_Message".tALM.tW);

   END_IF;
END_REGION

